(* Logix 5000 project; controller MV vendor 1 type 14 code 217 rev 31.11; software revision 31.00; part 44 of 53 *)
(* tags used below, declared in another part *)
   Always_Off : BOOL;
   CWD : CHECKWORD_FLAGS;
   MC_N100 : INT[255];   // C1_PLC Channel 1 PLC data
   MC_N120 : INT[255];   // C2 PLC Channel 2 PLC data
   MV21_TP_Capture_Volume_Timer : TIMER;
   MV_BM01_AV01_CIP : BOOL;
   MV_BM01_ZS04 : PlantItem;   // BM01ZS04
   MV_BM01_ZS05 : PlantItem;   // BM01ZS05
   MV_Data_To_TF : DINT[30];
   MV_Enable_MV21_NewPressureControl : BOOL;
   MV_FP01_ZS01 : PlantItem;   // FP01ZS01
   MV_FP01_ZS02 : PlantItem;   // FP01ZS02
   MV_MV20_CIP : BOOL;
   MV_MV20_TP_Command : DINT;
   MV_MV20_TP_Faulted : BOOL;
   MV_MV20_TP_Held : BOOL;
   MV_MV20_TP_NotIdle : BOOL;
   MV_MV20_TP_Prompt : DINT;
   MV_MV20_TP_Running : BOOL;
   MV_MV20_TP_Status : DINT;   // 0 = Idle, 1 = Running, 2 = Held, 3 = Faulted
   MV_MV20_TP_Step : DINT;
   MV_MV21_CO2_ON_PreStorage : BOOL;
   MV_MV21_CO2_ON_Storage : BOOL;
   MV_MV21_Filling_PulseLevel : REAL;
   MV_MV21_LTX07_TrueLevel : REAL;
   MV_MV21_ProxiesOK : BOOL;
   MV_MV21_PTX01_AI : PlantItem;   // MV21_PTX01
   MV_MV21_TP_CaskDepressure : BOOL;
   MV_MV21_TP_CaskEmptying : BOOL;
   MV_MV21_TP_CaskFilling : BOOL;
   MV_MV21_TP_CaskPreEmptyPressure : BOOL;
   MV_MV21_TP_CaskPrePressure : BOOL;
   MV_MV21_TP_CaskPressureDelay : BOOL;
   MV_MV21_TP_CaskPurgeFromTop : BOOL;
   MV_MV21_TP_CaskReadyToFill : BOOL;
   MV_MV21_TP_CaskStorage : BOOL;
   MV_MV21_TP_Command : DINT;
   MV_MV21_TP_DAL_Chase_Cask : BOOL;
   MV_MV21_TP_DAL_Chase_KB : BOOL;
   MV_MV21_TP_DAL_Chase_Time : TIMER;
   MV_MV21_TP_Dirty : BOOL;
   MV_MV21_TP_Emptying_Level_Setpoint : REAL;
   MV_MV21_TP_Error_String : STRING;
   MV_MV21_TP_Idle : BOOL;
   MV_MV21_TP_Initial_DAL_Chase_Cask : BOOL;
   MV_MV21_TP_Initial_DAL_Chase_KB : BOOL;
   MV_MV21_TP_KBDepressure : BOOL;
   MV_MV21_TP_KBEmptying : BOOL;
   MV_MV21_TP_KBFilling : BOOL;
   MV_MV21_TP_KBFilling_M : BOOL;
   MV_MV21_TP_KBPreEmptyPressure : BOOL;
   MV_MV21_TP_KBPrePressurise : BOOL;
   MV_MV21_TP_KBPurgeFromTop : BOOL;
   MV_MV21_TP_KBPurgeTimer : TIMER;
   MV_MV21_TP_KBStorage : BOOL;
   MV_MV21_TP_LowerLimit : REAL;
   MV_MV21_TP_ONS : BOOL;
   MV_MV21_TP_ONS_1 : BOOL;
   MV_MV21_TP_Prompt : DINT;
   MV_MV21_TP_Proxy_Delay_Made : TIMER;
   MV_MV21_TP_Proxy_Delay_NOT_MADE : TIMER;
   MV_MV21_TP_ReadyToFillKB : BOOL;
   MV_MV21_TP_ReadyToFillKB_M : BOOL;
   MV_MV21_TP_Running : BOOL;
   MV_MV21_TP_Setpoint : REAL;
   MV_MV21_TP_Status : DINT;   // 0 = Idle, 1 = Running, 2 = Held, 3 = Faulted
   MV_MV21_TP_Step : DINT;
   MV_MV21_TP_Steptime : DINT;
   MV_MV21_TP_UpperLimit : REAL;
   MV_MV21_TP_Vent : BOOL;
   MV_MV21_Transfer_StartLevel : REAL;
   MV_MV21_Transferred_Level : REAL;
   MV_N137 : INT[50];   // MV 21, CURRENT FV DATA
   MV_TP_CaskEmptyingPressure : REAL;
   MV_TP_CaskFillingPressure : REAL;
   MV_TP_CaskPrefillPressure : REAL;
   MV_TP_CaskStoragePressure : REAL;
   MV_TP_CaskStoragePressureDelay : DINT;
   MV_TP_CaskStoragePressureDelay_Secs : DINT;
   MV_TP_CaskStoragePressureLevel : REAL;
   MV_TP_Emptying_Volume_Setpoint : REAL;
   MV_TP_KBEmptyingPressure : REAL;
   MV_TP_KBFillingPressure : REAL;
   MV_TP_KBPrefillPressure : REAL;
   MV_TP_KBStoragePressure : REAL;
   MV_TP_KBStoragePressureLevel : REAL;
   MV_TP_NoCIPDelay : DINT;
   MV_TP_VentPressure : REAL;
(* MV_Common, continued *)

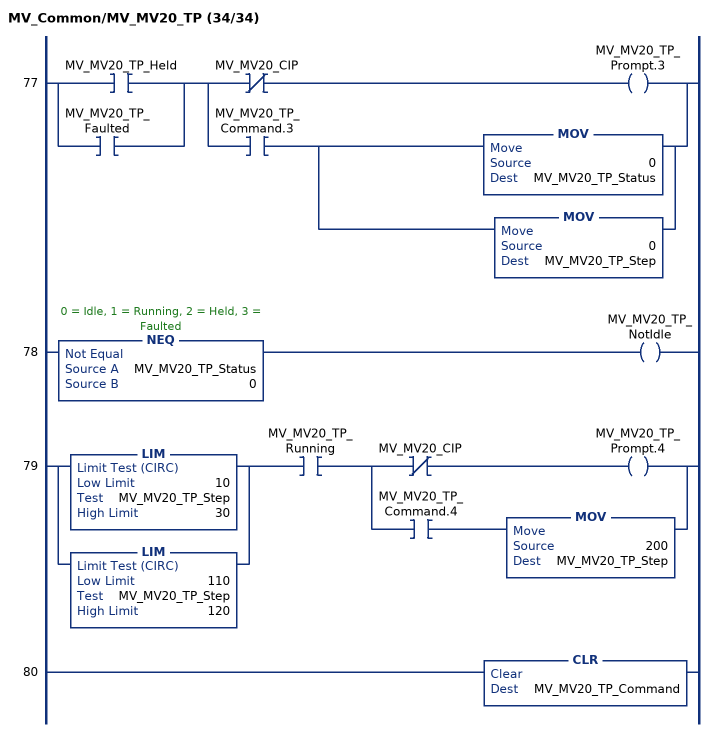
   77: [XIC(MV_MV20_TP_Held) ,XIC(MV_MV20_TP_Faulted) ][XIO(MV_MV20_CIP) OTE(MV_MV20_TP_Prompt.3) ,XIC(MV_MV20_TP_Command.3) [MOV(0,MV_MV20_TP_Status) ,MOV(0,MV_MV20_TP_Step) ] ];
   78: NEQ(MV_MV20_TP_Status,0)OTE(MV_MV20_TP_NotIdle);
   79: [LIM(10,MV_MV20_TP_Step,30) ,LIM(110,MV_MV20_TP_Step,120) ]XIC(MV_MV20_TP_Running)[XIO(MV_MV20_CIP) OTE(MV_MV20_TP_Prompt.4) ,XIC(MV_MV20_TP_Command.4) MOV(200,MV_MV20_TP_Step) ];
   80: CLR(MV_MV20_TP_Command);
END_ROUTINE

ROUTINE MV_MV21_TP   (* ladder *)
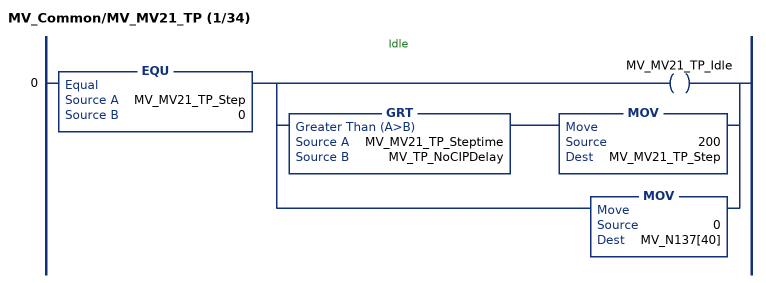
   // Idle
   0: EQU(MV_MV21_TP_Step,0)[OTE(MV_MV21_TP_Idle) ,GRT(MV_MV21_TP_Steptime,MV_TP_NoCIPDelay) MOV(200,MV_MV21_TP_Step) ,MOV(0,MV_N137[40]) ];
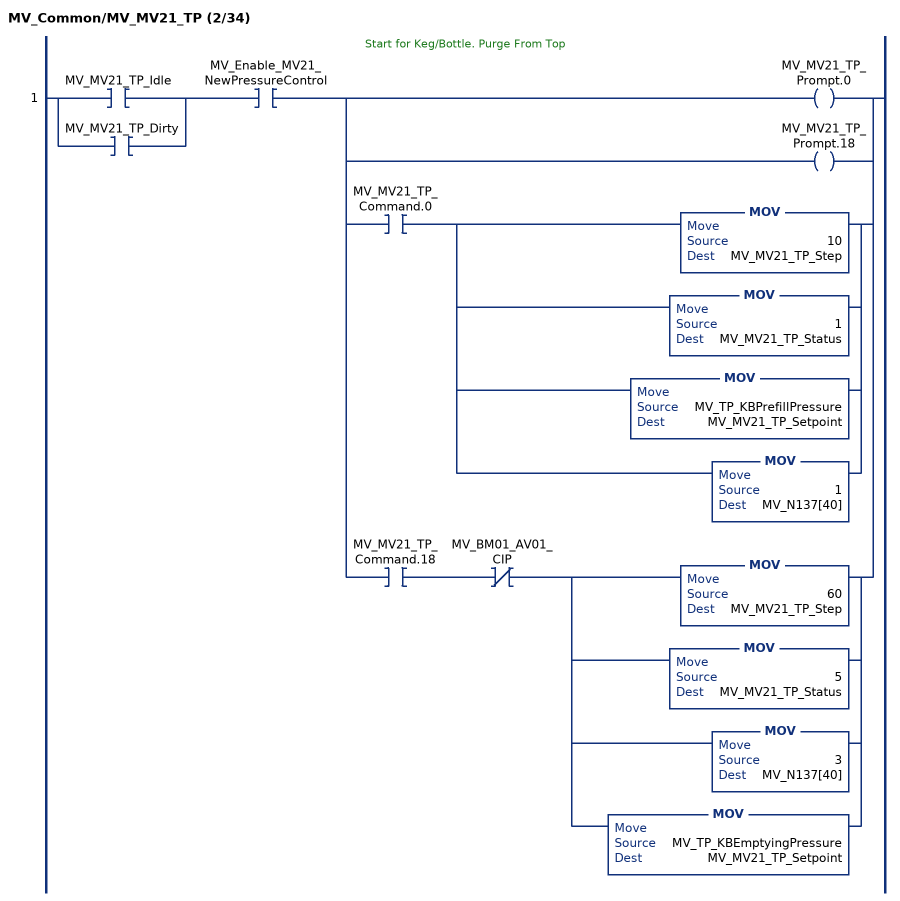
   // Start for Keg/Bottle. Purge From Top
   1: [XIC(MV_MV21_TP_Idle) ,XIC(MV_MV21_TP_Dirty) ]XIC(MV_Enable_MV21_NewPressureControl)[OTE(MV_MV21_TP_Prompt.0) ,OTE(MV_MV21_TP_Prompt.18) ,XIC(MV_MV21_TP_Command.0) [MOV(10,MV_MV21_TP_Step) ,MOV(1,MV_MV21_TP_Status) ,MOV(MV_TP_KBPrefillPressure,MV_MV21_TP_Setpoint) ,MOV(1,MV_N137[40]) ] ,XIC(MV_MV21_TP_Command.18) XIO(MV_BM01_AV01_CIP) [MOV(60,MV_MV21_TP_Step) ,MOV(5,MV_MV21_TP_Status) ,MOV(3,MV_N137[40]) ,MOV(MV_TP_KBEmptyingPressure,MV_MV21_TP_Setpoint) ] ];
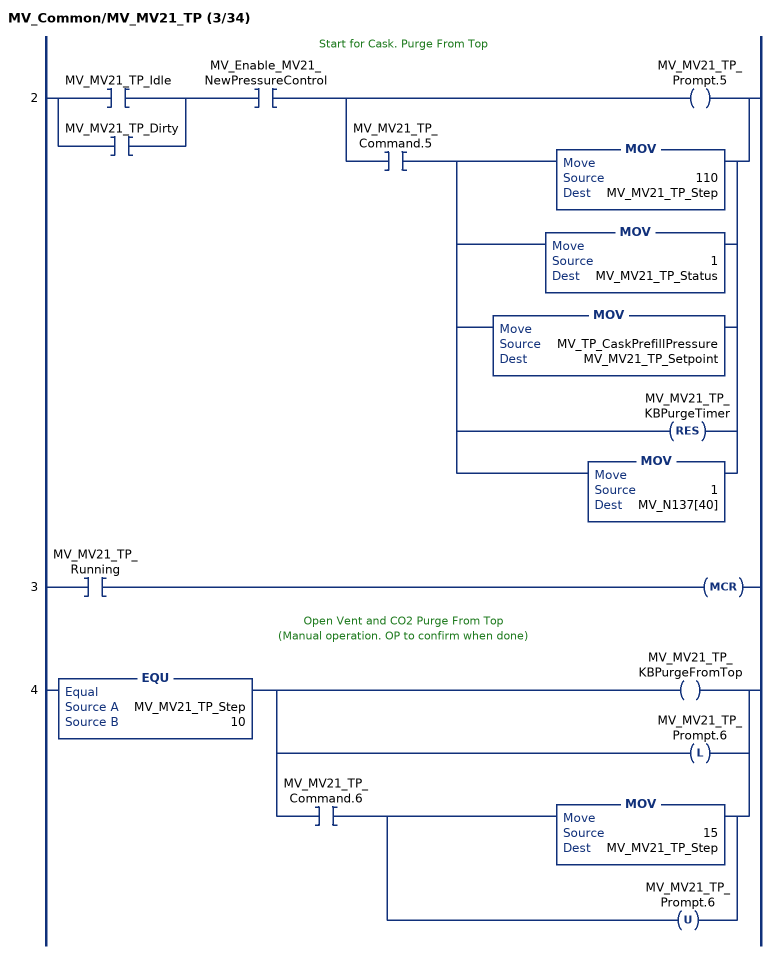
   // Start for Cask. Purge From Top
   2: [XIC(MV_MV21_TP_Idle) ,XIC(MV_MV21_TP_Dirty) ]XIC(MV_Enable_MV21_NewPressureControl)[OTE(MV_MV21_TP_Prompt.5) ,XIC(MV_MV21_TP_Command.5) [MOV(110,MV_MV21_TP_Step) ,MOV(1,MV_MV21_TP_Status) ,MOV(MV_TP_CaskPrefillPressure,MV_MV21_TP_Setpoint) ,RES(MV_MV21_TP_KBPurgeTimer) ,MOV(1,MV_N137[40]) ] ];
   3: XIC(MV_MV21_TP_Running)MCR();
   // Open Vent and CO2 Purge From Top
   // (Manual operation. OP to confirm when done)
   4: EQU(MV_MV21_TP_Step,10)[OTE(MV_MV21_TP_KBPurgeFromTop) ,OTL(MV_MV21_TP_Prompt.6) ,XIC(MV_MV21_TP_Command.6) [MOV(15,MV_MV21_TP_Step) ,OTU(MV_MV21_TP_Prompt.6) ] ];
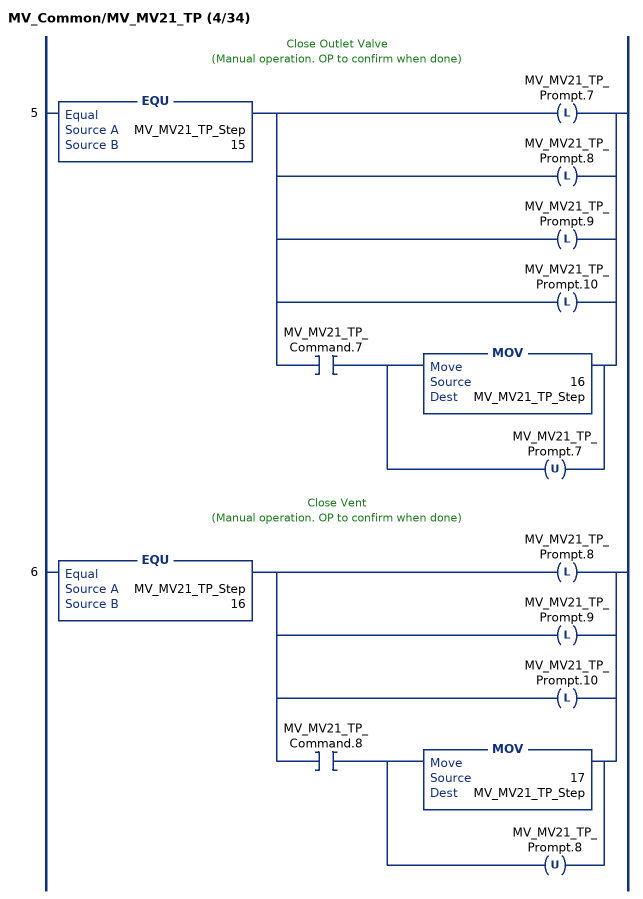
   // Close Outlet Valve
   // (Manual operation. OP to confirm when done)
   5: EQU(MV_MV21_TP_Step,15)[OTL(MV_MV21_TP_Prompt.7) ,OTL(MV_MV21_TP_Prompt.8) ,OTL(MV_MV21_TP_Prompt.9) ,OTL(MV_MV21_TP_Prompt.10) ,XIC(MV_MV21_TP_Command.7) [MOV(16,MV_MV21_TP_Step) ,OTU(MV_MV21_TP_Prompt.7) ] ];
   // Close Vent
   // (Manual operation. OP to confirm when done)
   6: EQU(MV_MV21_TP_Step,16)[OTL(MV_MV21_TP_Prompt.8) ,OTL(MV_MV21_TP_Prompt.9) ,OTL(MV_MV21_TP_Prompt.10) ,XIC(MV_MV21_TP_Command.8) [MOV(17,MV_MV21_TP_Step) ,OTU(MV_MV21_TP_Prompt.8) ] ];
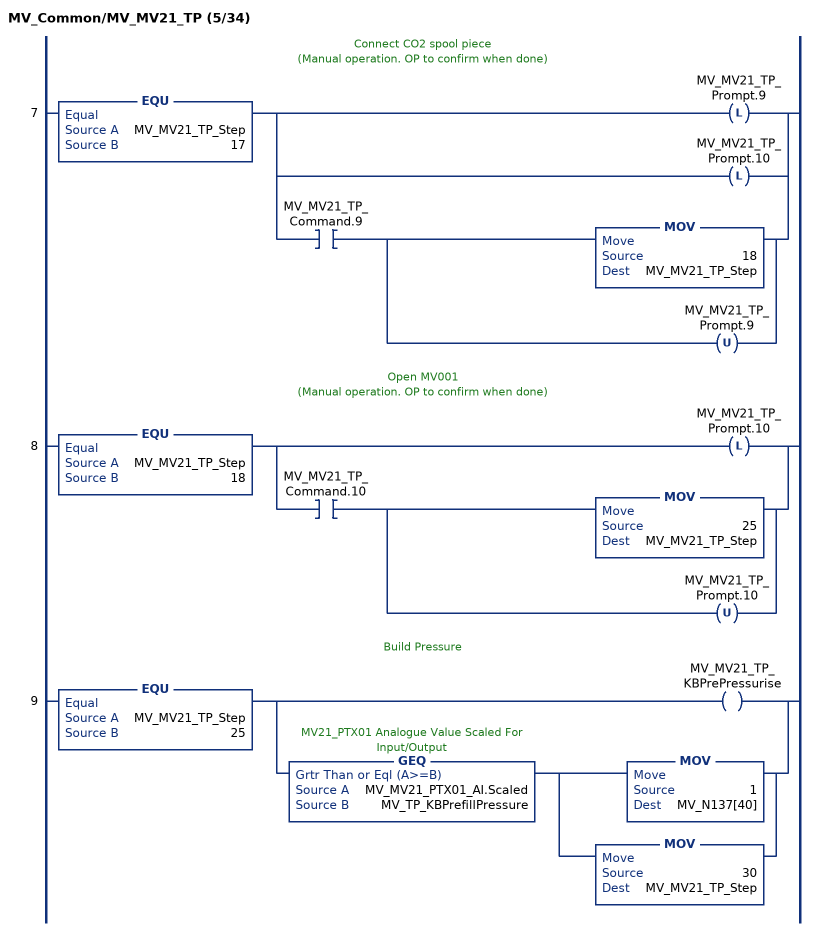
   // Connect CO2 spool piece
   // (Manual operation. OP to confirm when done)
   7: EQU(MV_MV21_TP_Step,17)[OTL(MV_MV21_TP_Prompt.9) ,OTL(MV_MV21_TP_Prompt.10) ,XIC(MV_MV21_TP_Command.9) [MOV(18,MV_MV21_TP_Step) ,OTU(MV_MV21_TP_Prompt.9) ] ];
   // Open MV001
   // (Manual operation. OP to confirm when done)
   8: EQU(MV_MV21_TP_Step,18)[OTL(MV_MV21_TP_Prompt.10) ,XIC(MV_MV21_TP_Command.10) [MOV(25,MV_MV21_TP_Step) ,OTU(MV_MV21_TP_Prompt.10) ] ];
   // Build Pressure
   9: EQU(MV_MV21_TP_Step,25)[OTE(MV_MV21_TP_KBPrePressurise) ,GEQ(MV_MV21_PTX01_AI.Scaled,MV_TP_KBPrefillPressure) [MOV(1,MV_N137[40]) ,MOV(30,MV_MV21_TP_Step) ] ];
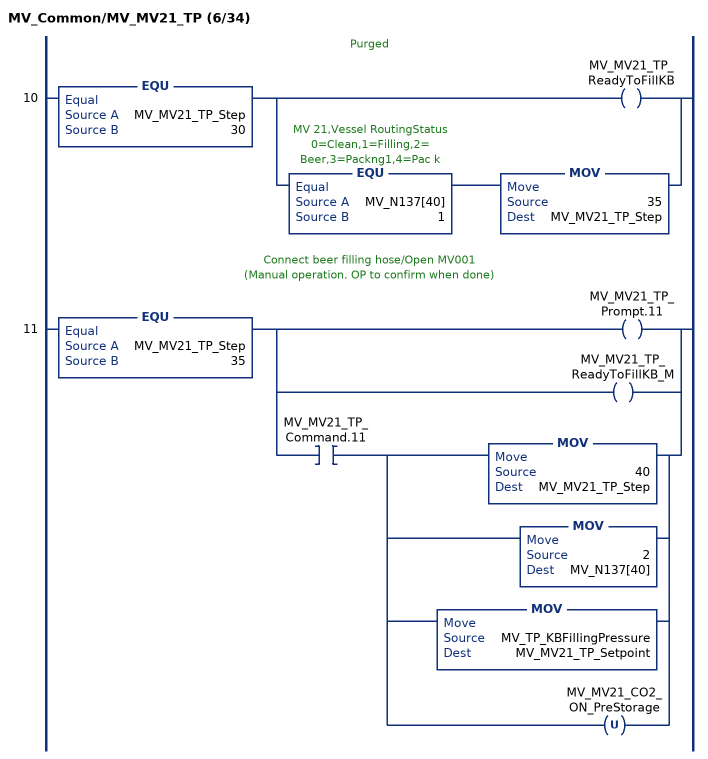
   // Purged
   10: EQU(MV_MV21_TP_Step,30)[OTE(MV_MV21_TP_ReadyToFillKB) ,EQU(MV_N137[40],1) MOV(35,MV_MV21_TP_Step) ];
   // Connect beer filling hose/Open MV001
   // (Manual operation. OP to confirm when done)
   11: EQU(MV_MV21_TP_Step,35)[OTE(MV_MV21_TP_Prompt.11) ,OTE(MV_MV21_TP_ReadyToFillKB_M) ,XIC(MV_MV21_TP_Command.11) [MOV(40,MV_MV21_TP_Step) ,MOV(2,MV_N137[40]) ,MOV(MV_TP_KBFillingPressure,MV_MV21_TP_Setpoint) ,OTU(MV_MV21_CO2_ON_PreStorage) ] ];
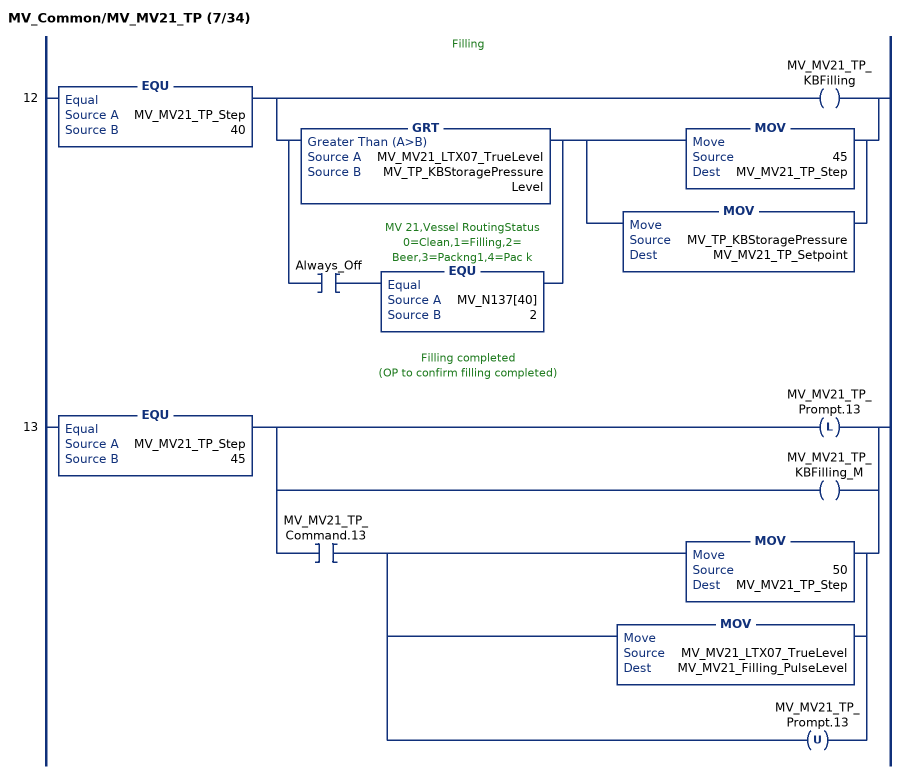
   // Filling
   12: EQU(MV_MV21_TP_Step,40)[OTE(MV_MV21_TP_KBFilling) ,[GRT(MV_MV21_LTX07_TrueLevel,MV_TP_KBStoragePressureLevel) ,XIC(Always_Off) EQU(MV_N137[40],2) ] [MOV(45,MV_MV21_TP_Step) ,MOV(MV_TP_KBStoragePressure,MV_MV21_TP_Setpoint) ] ];
   // Filling completed
   // (OP to confirm filling completed)
   13: EQU(MV_MV21_TP_Step,45)[OTL(MV_MV21_TP_Prompt.13) ,OTE(MV_MV21_TP_KBFilling_M) ,XIC(MV_MV21_TP_Command.13) [MOV(50,MV_MV21_TP_Step) ,MOV(MV_MV21_LTX07_TrueLevel,MV_MV21_Filling_PulseLevel) ,OTU(MV_MV21_TP_Prompt.13) ] ];
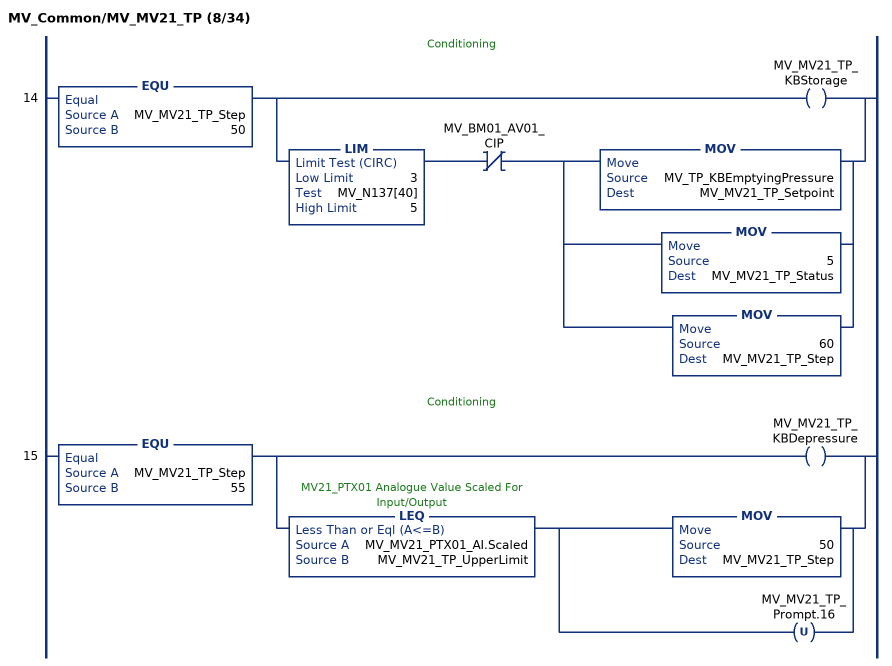
   // Conditioning
   14: EQU(MV_MV21_TP_Step,50)[OTE(MV_MV21_TP_KBStorage) ,LIM(3,MV_N137[40],5) XIO(MV_BM01_AV01_CIP) [MOV(MV_TP_KBEmptyingPressure,MV_MV21_TP_Setpoint) ,MOV(5,MV_MV21_TP_Status) ,MOV(60,MV_MV21_TP_Step) ] ];
   // Conditioning
   15: EQU(MV_MV21_TP_Step,55)[OTE(MV_MV21_TP_KBDepressure) ,LEQ(MV_MV21_PTX01_AI.Scaled,MV_MV21_TP_UpperLimit) [MOV(50,MV_MV21_TP_Step) ,OTU(MV_MV21_TP_Prompt.16) ] ];
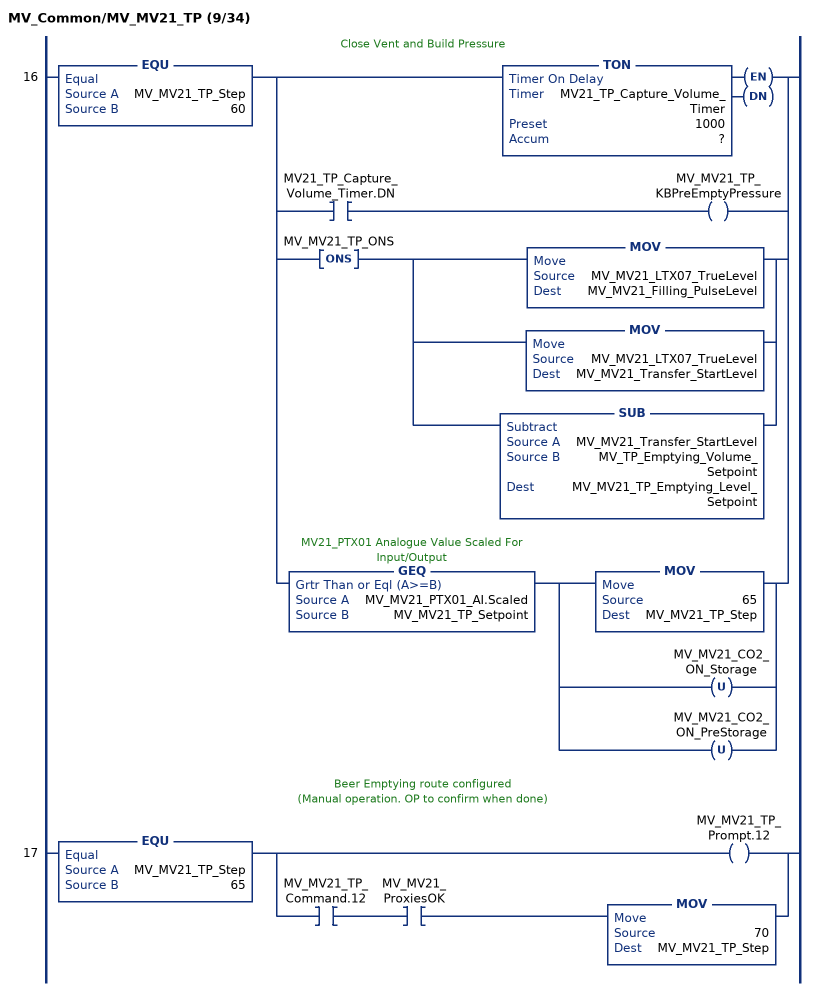
   // Close Vent and Build Pressure
   16: EQU(MV_MV21_TP_Step,60)[TON(MV21_TP_Capture_Volume_Timer,?,?) ,XIC(MV21_TP_Capture_Volume_Timer.DN) OTE(MV_MV21_TP_KBPreEmptyPressure) ,ONS(MV_MV21_TP_ONS) [MOV(MV_MV21_LTX07_TrueLevel,MV_MV21_Filling_PulseLevel) ,MOV(MV_MV21_LTX07_TrueLevel,MV_MV21_Transfer_StartLevel) ,SUB(MV_MV21_Transfer_StartLevel,MV_TP_Emptying_Volume_Setpoint,MV_MV21_TP_Emptying_Level_Setpoint) ] ,GEQ(MV_MV21_PTX01_AI.Scaled,MV_MV21_TP_Setpoint) [MOV(65,MV_MV21_TP_Step) ,OTU(MV_MV21_CO2_ON_Storage) ,OTU(MV_MV21_CO2_ON_PreStorage) ] ];
   // Beer Emptying route configured
   // (Manual operation. OP to confirm when done)
   17: EQU(MV_MV21_TP_Step,65)[OTE(MV_MV21_TP_Prompt.12) ,XIC(MV_MV21_TP_Command.12) XIC(MV_MV21_ProxiesOK) MOV(70,MV_MV21_TP_Step) ];
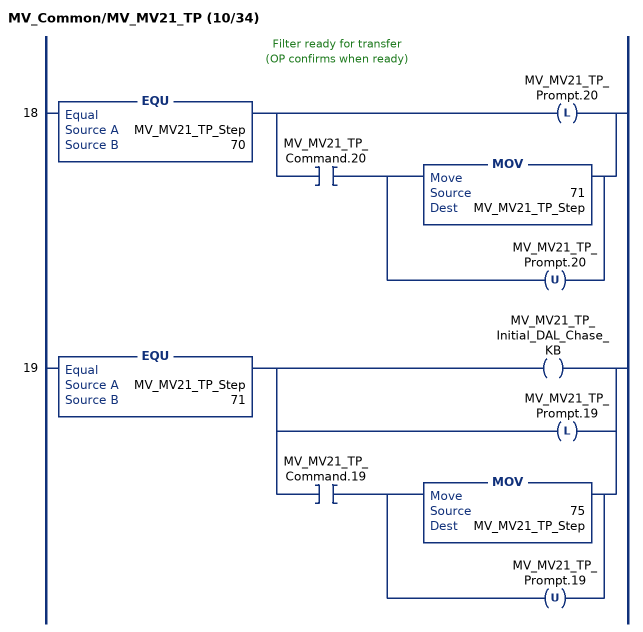
   // Filter ready for transfer
   // (OP confirms when ready)
   18: EQU(MV_MV21_TP_Step,70)[OTL(MV_MV21_TP_Prompt.20) ,XIC(MV_MV21_TP_Command.20) [MOV(71,MV_MV21_TP_Step) ,OTU(MV_MV21_TP_Prompt.20) ] ];
   19: EQU(MV_MV21_TP_Step,71)[OTE(MV_MV21_TP_Initial_DAL_Chase_KB) ,OTL(MV_MV21_TP_Prompt.19) ,XIC(MV_MV21_TP_Command.19) [MOV(75,MV_MV21_TP_Step) ,OTU(MV_MV21_TP_Prompt.19) ] ];